   // stn[3].wipBtn[49,6] := 1000;
   // stn[3].wipBtn[49,7] := 1000;
   // stn[4].wipBtn[0,0] := 1000;
   // stn[4].wipBtn[0,1] := 1000;
   // stn[4].wipBtn[0,2] := 1000;
   // stn[4].wipBtn[0,3] := 1000;
   // stn[4].wipBtn[0,4] := 1000;
   // stn[4].wipBtn[0,5] := 1000;
   // stn[4].wipBtn[0,6] := 1000;
   // stn[4].wipBtn[0,7] := 195000;
   // stn[4].wipBtn[1,0] := 1000;
   // stn[4].wipBtn[1,1] := 1000;
   // stn[4].wipBtn[1,2] := 1000;
   // stn[4].wipBtn[1,3] := 1000;
   // stn[4].wipBtn[1,4] := 1000;
   // stn[4].wipBtn[1,5] := 1000;
   // stn[4].wipBtn[1,6] := 1000;
   // stn[4].wipBtn[1,7] := 1000;
   // stn[4].wipBtn[2,0] := 1000;
   // stn[4].wipBtn[2,1] := 1000;
   // stn[4].wipBtn[2,2] := 1000;
   // stn[4].wipBtn[2,3] := 1000;
   // stn[4].wipBtn[2,4] := 1000;
   // stn[4].wipBtn[2,5] := 1000;
   // stn[4].wipBtn[2,6] := 1000;
   // stn[4].wipBtn[2,7] := 1000;
   // stn[4].wipBtn[3,0] := 1000;
   // stn[4].wipBtn[3,1] := 1000;
   // stn[4].wipBtn[3,2] := 1000;
   // stn[4].wipBtn[3,3] := 1000;
   // stn[4].wipBtn[3,4] := 1000;
   // stn[4].wipBtn[3,5] := 1000;
   // stn[4].wipBtn[3,6] := 1000;
   // stn[4].wipBtn[3,7] := 1000;
   // stn[4].wipBtn[4,0] := 1000;
   // stn[4].wipBtn[4,1] := 1000;
   // stn[4].wipBtn[4,2] := 1000;
   // stn[4].wipBtn[4,3] := 1000;
   // stn[4].wipBtn[4,4] := 1000;
   // stn[4].wipBtn[4,5] := 1000;
   // stn[4].wipBtn[4,6] := 1000;
   // stn[4].wipBtn[4,7] := 1000;
   // stn[4].wipBtn[5,0] := 1000;
   // stn[4].wipBtn[5,1] := 1000;
   // stn[4].wipBtn[5,2] := 1000;
   // stn[4].wipBtn[5,3] := 1000;
   // stn[4].wipBtn[5,4] := 1000;
   // stn[4].wipBtn[5,5] := 1000;
   // stn[4].wipBtn[5,6] := 1000;
   // stn[4].wipBtn[5,7] := 1000;
   // stn[4].wipBtn[6,0] := 1000;
   // stn[4].wipBtn[6,1] := 1000;
   // stn[4].wipBtn[6,2] := 1000;
   // stn[4].wipBtn[6,3] := 1000;
   // stn[4].wipBtn[6,4] := 1000;
   // stn[4].wipBtn[6,5] := 1000;
   // stn[4].wipBtn[6,6] := 1000;
   // stn[4].wipBtn[6,7] := 1000;
   // stn[4].wipBtn[7,0] := 1000;
   // stn[4].wipBtn[7,1] := 1000;
   // stn[4].wipBtn[7,2] := 1000;
   // stn[4].wipBtn[7,3] := 1000;
   // stn[4].wipBtn[7,4] := 1000;
   // stn[4].wipBtn[7,5] := 1000;
   // stn[4].wipBtn[7,6] := 1000;
   // stn[4].wipBtn[7,7] := 1000;
   // stn[4].wipBtn[8,0] := 1000;
   // stn[4].wipBtn[8,1] := 1000;
   // stn[4].wipBtn[8,2] := 1000;
   // stn[4].wipBtn[8,3] := 1000;
   // stn[4].wipBtn[8,4] := 1000;
   // stn[4].wipBtn[8,5] := 1000;
   // stn[4].wipBtn[8,6] := 1000;
   // stn[4].wipBtn[8,7] := 1000;
   // stn[4].wipBtn[9,0] := 1000;
   // stn[4].wipBtn[9,1] := 1000;
   // stn[4].wipBtn[9,2] := 1000;
   // stn[4].wipBtn[9,3] := 1000;
   // stn[4].wipBtn[9,4] := 1000;
   // stn[4].wipBtn[9,5] := 1000;
   // stn[4].wipBtn[9,6] := 1000;
   // stn[4].wipBtn[9,7] := 1000;
   // stn[4].wipBtn[10,0] := 1000;
   // stn[4].wipBtn[10,1] := 1000;
   // stn[4].wipBtn[10,2] := 1000;
   // stn[4].wipBtn[10,3] := 1000;
   // stn[4].wipBtn[10,4] := 1000;
   // stn[4].wipBtn[10,5] := 1000;
   // stn[4].wipBtn[10,6] := 1000;
   // stn[4].wipBtn[10,7] := 1000;
   // stn[4].wipBtn[11,0] := 1000;
   // stn[4].wipBtn[11,1] := 1000;
   // stn[4].wipBtn[11,2] := 1000;
   // stn[4].wipBtn[11,3] := 1000;
   // stn[4].wipBtn[11,4] := 1000;
   // stn[4].wipBtn[11,5] := 1000;
   // stn[4].wipBtn[11,6] := 1000;
   // stn[4].wipBtn[11,7] := 1000;
   // stn[4].wipBtn[12,0] := 1000;
   // stn[4].wipBtn[12,1] := 1000;
   // stn[4].wipBtn[12,2] := 1000;
   // stn[4].wipBtn[12,3] := 1000;
   // stn[4].wipBtn[12,4] := 1000;
   // stn[4].wipBtn[12,5] := 1000;
   // stn[4].wipBtn[12,6] := 1000;
   // stn[4].wipBtn[12,7] := 1000;
   // stn[4].wipBtn[13,0] := 1000;
   // stn[4].wipBtn[13,1] := 1000;
   // stn[4].wipBtn[13,2] := 1000;
   // stn[4].wipBtn[13,3] := 1000;
   // stn[4].wipBtn[13,4] := 1000;
   // stn[4].wipBtn[13,5] := 1000;
   // stn[4].wipBtn[13,6] := 1000;
   // stn[4].wipBtn[13,7] := 1000;
   // stn[4].wipBtn[14,0] := 1000;
   // stn[4].wipBtn[14,1] := 1000;
   // stn[4].wipBtn[14,2] := 1000;
   // stn[4].wipBtn[14,3] := 1000;
   // stn[4].wipBtn[14,4] := 1000;
   // stn[4].wipBtn[14,5] := 1000;
   // stn[4].wipBtn[14,6] := 1000;
   // stn[4].wipBtn[14,7] := 1000;
   // stn[4].wipBtn[15,0] := 1000;
   // stn[4].wipBtn[15,1] := 1000;
   // stn[4].wipBtn[15,2] := 1000;
   // stn[4].wipBtn[15,3] := 1000;
   // stn[4].wipBtn[15,4] := 1000;
   // stn[4].wipBtn[15,5] := 1000;
   // stn[4].wipBtn[15,6] := 1000;
   // stn[4].wipBtn[15,7] := 1000;
   // stn[4].wipBtn[16,0] := 1000;
   // stn[4].wipBtn[16,1] := 1000;
   // stn[4].wipBtn[16,2] := 1000;
   // stn[4].wipBtn[16,3] := 1000;
   // stn[4].wipBtn[16,4] := 1000;
   // stn[4].wipBtn[16,5] := 1000;
   // stn[4].wipBtn[16,6] := 1000;
   // stn[4].wipBtn[16,7] := 1000;
   // stn[4].wipBtn[17,0] := 1000;
   // stn[4].wipBtn[17,1] := 1000;
   // stn[4].wipBtn[17,2] := 1000;
   // stn[4].wipBtn[17,3] := 1000;
   // stn[4].wipBtn[17,4] := 1000;
   // stn[4].wipBtn[17,5] := 1000;
   // stn[4].wipBtn[17,6] := 1000;
   // stn[4].wipBtn[17,7] := 1000;
   // stn[4].wipBtn[18,0] := 1000;
   // stn[4].wipBtn[18,1] := 1000;
   // stn[4].wipBtn[18,2] := 1000;
   // stn[4].wipBtn[18,3] := 1000;
   // stn[4].wipBtn[18,4] := 1000;
   // stn[4].wipBtn[18,5] := 1000;
   // stn[4].wipBtn[18,6] := 1000;
   // stn[4].wipBtn[18,7] := 1000;
   // stn[4].wipBtn[19,0] := 1000;
   // stn[4].wipBtn[19,1] := 1000;
   // stn[4].wipBtn[19,2] := 1000;
   // stn[4].wipBtn[19,3] := 1000;
   // stn[4].wipBtn[19,4] := 1000;
   // stn[4].wipBtn[19,5] := 1000;
   // stn[4].wipBtn[19,6] := 1000;
   // stn[4].wipBtn[19,7] := 1000;
   // stn[4].wipBtn[20,0] := 1000;
   // stn[4].wipBtn[20,1] := 1000;
   // stn[4].wipBtn[20,2] := 1000;
   // stn[4].wipBtn[20,3] := 1000;
   // stn[4].wipBtn[20,4] := 1000;
   // stn[4].wipBtn[20,5] := 1000;
   // stn[4].wipBtn[20,6] := 1000;
   // stn[4].wipBtn[20,7] := 1000;
   // stn[4].wipBtn[21,0] := 1000;
   // stn[4].wipBtn[21,1] := 1000;
   // stn[4].wipBtn[21,2] := 1000;
   // stn[4].wipBtn[21,3] := 1000;
   // stn[4].wipBtn[21,4] := 1000;
   // stn[4].wipBtn[21,5] := 1000;
   // stn[4].wipBtn[21,6] := 1000;
   // stn[4].wipBtn[21,7] := 1000;
   // stn[4].wipBtn[22,0] := 1000;
   // stn[4].wipBtn[22,1] := 1000;
   // stn[4].wipBtn[22,2] := 1000;
   // stn[4].wipBtn[22,3] := 1000;
   // stn[4].wipBtn[22,4] := 1000;
   // stn[4].wipBtn[22,5] := 1000;
   // stn[4].wipBtn[22,6] := 1000;
   // stn[4].wipBtn[22,7] := 1000;
   // stn[4].wipBtn[23,0] := 1000;
   // stn[4].wipBtn[23,1] := 1000;
   // stn[4].wipBtn[23,2] := 1000;
   // stn[4].wipBtn[23,3] := 1000;
   // stn[4].wipBtn[23,4] := 1000;
   // stn[4].wipBtn[23,5] := 1000;
   // stn[4].wipBtn[23,6] := 1000;
   // stn[4].wipBtn[23,7] := 1000;
   // stn[4].wipBtn[24,0] := 1000;
   // stn[4].wipBtn[24,1] := 1000;
   // stn[4].wipBtn[24,2] := 1000;
   // stn[4].wipBtn[24,3] := 1000;
   // stn[4].wipBtn[24,4] := 1000;
   // stn[4].wipBtn[24,5] := 1000;
   // stn[4].wipBtn[24,6] := 1000;
   // stn[4].wipBtn[24,7] := 1000;
   // stn[4].wipBtn[25,0] := 1000;
   // stn[4].wipBtn[25,1] := 1000;
   // stn[4].wipBtn[25,2] := 1000;
   // stn[4].wipBtn[25,3] := 1000;
   // stn[4].wipBtn[25,4] := 1000;
   // stn[4].wipBtn[25,5] := 1000;
   // stn[4].wipBtn[25,6] := 1000;
   // stn[4].wipBtn[25,7] := 1000;
   // stn[4].wipBtn[26,0] := 1000;
   // stn[4].wipBtn[26,1] := 1000;
   // stn[4].wipBtn[26,2] := 1000;
   // stn[4].wipBtn[26,3] := 1000;
   // stn[4].wipBtn[26,4] := 1000;
   // stn[4].wipBtn[26,5] := 1000;
   // stn[4].wipBtn[26,6] := 1000;
   // stn[4].wipBtn[26,7] := 1000;
   // stn[4].wipBtn[27,0] := 1000;
   // stn[4].wipBtn[27,1] := 1000;
   // stn[4].wipBtn[27,2] := 1000;
   // stn[4].wipBtn[27,3] := 1000;
   // stn[4].wipBtn[27,4] := 1000;
   // stn[4].wipBtn[27,5] := 1000;
   // stn[4].wipBtn[27,6] := 1000;
   // stn[4].wipBtn[27,7] := 1000;
   // stn[4].wipBtn[28,0] := 1000;
   // stn[4].wipBtn[28,1] := 1000;
   // stn[4].wipBtn[28,2] := 1000;
   // stn[4].wipBtn[28,3] := 1000;
   // stn[4].wipBtn[28,4] := 1000;
   // stn[4].wipBtn[28,5] := 1000;
   // stn[4].wipBtn[28,6] := 1000;
   // stn[4].wipBtn[28,7] := 1000;
   // stn[4].wipBtn[29,0] := 1000;
   // stn[4].wipBtn[29,1] := 1000;
   // stn[4].wipBtn[29,2] := 1000;
   // stn[4].wipBtn[29,3] := 1000;
   // stn[4].wipBtn[29,4] := 1000;
   // stn[4].wipBtn[29,5] := 1000;
   // stn[4].wipBtn[29,6] := 1000;
   // stn[4].wipBtn[29,7] := 1000;
   // stn[4].wipBtn[30,0] := 1000;
   // stn[4].wipBtn[30,1] := 1000;
   // stn[4].wipBtn[30,2] := 1000;
   // stn[4].wipBtn[30,3] := 1000;
   // stn[4].wipBtn[30,4] := 1000;
   // stn[4].wipBtn[30,5] := 1000;
   // stn[4].wipBtn[30,6] := 1000;
   // stn[4].wipBtn[30,7] := 1000;
   // stn[4].wipBtn[31,0] := 1000;
   // stn[4].wipBtn[31,1] := 1000;
   // stn[4].wipBtn[31,2] := 1000;
   // stn[4].wipBtn[31,3] := 1000;
   // stn[4].wipBtn[31,4] := 1000;
   // stn[4].wipBtn[31,5] := 1000;
   // stn[4].wipBtn[31,6] := 1000;
   // stn[4].wipBtn[31,7] := 1000;
   // stn[4].wipBtn[32,0] := 1000;
   // stn[4].wipBtn[32,1] := 1000;
   // stn[4].wipBtn[32,2] := 1000;
   // stn[4].wipBtn[32,3] := 1000;
   // stn[4].wipBtn[32,4] := 1000;
   // stn[4].wipBtn[32,5] := 1000;
   // stn[4].wipBtn[32,6] := 1000;
   // stn[4].wipBtn[32,7] := 1000;
   // stn[4].wipBtn[33,0] := 1000;
   // stn[4].wipBtn[33,1] := 1000;
   // stn[4].wipBtn[33,2] := 1000;
   // stn[4].wipBtn[33,3] := 1000;
   // stn[4].wipBtn[33,4] := 1000;
   // stn[4].wipBtn[33,5] := 1000;
   // stn[4].wipBtn[33,6] := 1000;
   // stn[4].wipBtn[33,7] := 1000;
   // stn[4].wipBtn[34,0] := 1000;
   // stn[4].wipBtn[34,1] := 1000;
   // stn[4].wipBtn[34,2] := 1000;
   // stn[4].wipBtn[34,3] := 1000;
   // stn[4].wipBtn[34,4] := 1000;
   // stn[4].wipBtn[34,5] := 1000;
   // stn[4].wipBtn[34,6] := 1000;
   // stn[4].wipBtn[34,7] := 1000;
   // stn[4].wipBtn[35,0] := 1000;
   // stn[4].wipBtn[35,1] := 1000;
   // stn[4].wipBtn[35,2] := 1000;
   // stn[4].wipBtn[35,3] := 1000;
   // stn[4].wipBtn[35,4] := 1000;
   // stn[4].wipBtn[35,5] := 1000;
   // stn[4].wipBtn[35,6] := 1000;
   // stn[4].wipBtn[35,7] := 1000;
   // stn[4].wipBtn[36,0] := 1000;
   // stn[4].wipBtn[36,1] := 1000;
   // stn[4].wipBtn[36,2] := 1000;
   // stn[4].wipBtn[36,3] := 1000;
   // stn[4].wipBtn[36,4] := 1000;
   // stn[4].wipBtn[36,5] := 1000;
   // stn[4].wipBtn[36,6] := 1000;
   // stn[4].wipBtn[36,7] := 1000;
   // stn[4].wipBtn[37,0] := 1000;
   // stn[4].wipBtn[37,1] := 1000;
   // stn[4].wipBtn[37,2] := 1000;
   // stn[4].wipBtn[37,3] := 1000;
   // stn[4].wipBtn[37,4] := 1000;
   // stn[4].wipBtn[37,5] := 1000;
   // stn[4].wipBtn[37,6] := 1000;
   // stn[4].wipBtn[37,7] := 1000;
   // stn[4].wipBtn[38,0] := 1000;
   // stn[4].wipBtn[38,1] := 1000;
   // stn[4].wipBtn[38,2] := 1000;
   // stn[4].wipBtn[38,3] := 1000;
   // stn[4].wipBtn[38,4] := 1000;
   // stn[4].wipBtn[38,5] := 1000;
   // stn[4].wipBtn[38,6] := 1000;
   // stn[4].wipBtn[38,7] := 1000;
   // stn[4].wipBtn[39,0] := 1000;
   // stn[4].wipBtn[39,1] := 1000;
   // stn[4].wipBtn[39,2] := 1000;
   // stn[4].wipBtn[39,3] := 1000;
   // stn[4].wipBtn[39,4] := 1000;
   // stn[4].wipBtn[39,5] := 1000;
   // stn[4].wipBtn[39,6] := 1000;
   // stn[4].wipBtn[39,7] := 1000;
   // stn[4].wipBtn[40,0] := 1000;
   // stn[4].wipBtn[40,1] := 1000;
   // stn[4].wipBtn[40,2] := 1000;
   // stn[4].wipBtn[40,3] := 1000;
   // stn[4].wipBtn[40,4] := 1000;
   // stn[4].wipBtn[40,5] := 1000;
   // stn[4].wipBtn[40,6] := 1000;
   // stn[4].wipBtn[40,7] := 1000;
   // stn[4].wipBtn[41,0] := 1000;
   // stn[4].wipBtn[41,1] := 1000;
   // stn[4].wipBtn[41,2] := 1000;
   // stn[4].wipBtn[41,3] := 1000;
   // stn[4].wipBtn[41,4] := 1000;
   // stn[4].wipBtn[41,5] := 1000;
   // stn[4].wipBtn[41,6] := 1000;
   // stn[4].wipBtn[41,7] := 1000;
   // stn[4].wipBtn[42,0] := 1000;
   // stn[4].wipBtn[42,1] := 1000;
   // stn[4].wipBtn[42,2] := 1000;
   // stn[4].wipBtn[42,3] := 1000;
   // stn[4].wipBtn[42,4] := 1000;
   // stn[4].wipBtn[42,5] := 1000;
   // stn[4].wipBtn[42,6] := 1000;
   // stn[4].wipBtn[42,7] := 1000;
   // stn[4].wipBtn[43,0] := 1000;
   // stn[4].wipBtn[43,1] := 1000;
   // stn[4].wipBtn[43,2] := 1000;
   // stn[4].wipBtn[43,3] := 1000;
   // stn[4].wipBtn[43,4] := 1000;
   // stn[4].wipBtn[43,5] := 1000;
   // stn[4].wipBtn[43,6] := 1000;
   // stn[4].wipBtn[43,7] := 1000;
   // stn[4].wipBtn[44,0] := 1000;
   // stn[4].wipBtn[44,1] := 1000;
   // stn[4].wipBtn[44,2] := 1000;
   // stn[4].wipBtn[44,3] := 1000;
   // stn[4].wipBtn[44,4] := 1000;
   // stn[4].wipBtn[44,5] := 1000;
   // stn[4].wipBtn[44,6] := 1000;
   // stn[4].wipBtn[44,7] := 1000;
   // stn[4].wipBtn[45,0] := 1000;
   // stn[4].wipBtn[45,1] := 1000;
   // stn[4].wipBtn[45,2] := 1000;
   // stn[4].wipBtn[45,3] := 1000;
   // stn[4].wipBtn[45,4] := 1000;
   // stn[4].wipBtn[45,5] := 1000;
   // stn[4].wipBtn[45,6] := 1000;
   // stn[4].wipBtn[45,7] := 1000;
   // stn[4].wipBtn[46,0] := 1000;
   // stn[4].wipBtn[46,1] := 1000;
   // stn[4].wipBtn[46,2] := 1000;
   // stn[4].wipBtn[46,3] := 1000;
   // stn[4].wipBtn[46,4] := 1000;
   // stn[4].wipBtn[46,5] := 1000;
   // stn[4].wipBtn[46,6] := 1000;
   // stn[4].wipBtn[46,7] := 1000;
   // stn[4].wipBtn[47,0] := 1000;
   // stn[4].wipBtn[47,1] := 1000;
   // stn[4].wipBtn[47,2] := 1000;
   // stn[4].wipBtn[47,3] := 1000;
   // stn[4].wipBtn[47,4] := 1000;
   // stn[4].wipBtn[47,5] := 1000;
   // stn[4].wipBtn[47,6] := 1000;
   // stn[4].wipBtn[47,7] := 1000;
   // stn[4].wipBtn[48,0] := 1000;
   // stn[4].wipBtn[48,1] := 1000;
   // stn[4].wipBtn[48,2] := 1000;
   // stn[4].wipBtn[48,3] := 1000;
   // stn[4].wipBtn[48,4] := 1000;
   // stn[4].wipBtn[48,5] := 1000;
   // stn[4].wipBtn[48,6] := 1000;
   // stn[4].wipBtn[48,7] := 1000;
   // stn[4].wipBtn[49,0] := 1000;
   // stn[4].wipBtn[49,1] := 1000;
   // stn[4].wipBtn[49,2] := 1000;
   // stn[4].wipBtn[49,3] := 1000;
   // stn[4].wipBtn[49,4] := 1000;
   // stn[4].wipBtn[49,5] := 1000;
   // stn[4].wipBtn[49,6] := 1000;
   // stn[4].wipBtn[49,7] := 1000;
   // stn[5].wipBtn[0,0] := 1000;
   // stn[5].wipBtn[0,1] := 194000;
   // stn[5].wipBtn[0,2] := 196000;
   // stn[5].wipBtn[0,3] := 177000;
   // stn[5].wipBtn[0,4] := 1000;
   // stn[5].wipBtn[0,5] := 197000;
   // stn[5].wipBtn[0,6] := 178000;
   // stn[5].wipBtn[0,7] := 176000;
   // stn[5].wipBtn[1,0] := 1000;
   // stn[5].wipBtn[1,1] := 1000;
   // stn[5].wipBtn[1,2] := 1000;
   // stn[5].wipBtn[1,3] := 1000;
   // stn[5].wipBtn[1,4] := 1000;
   // stn[5].wipBtn[1,5] := 1000;
   // stn[5].wipBtn[1,6] := 1000;
   // stn[5].wipBtn[1,7] := 1000;
   // stn[5].wipBtn[2,0] := 1000;
   // stn[5].wipBtn[2,1] := 1000;
   // stn[5].wipBtn[2,2] := 1000;
   // stn[5].wipBtn[2,3] := 1000;
   // stn[5].wipBtn[2,4] := 1000;
   // stn[5].wipBtn[2,5] := 1000;
   // stn[5].wipBtn[2,6] := 1000;
   // stn[5].wipBtn[2,7] := 1000;
   // stn[5].wipBtn[3,0] := 1000;
   // stn[5].wipBtn[3,1] := 1000;
   // stn[5].wipBtn[3,2] := 1000;
   // stn[5].wipBtn[3,3] := 1000;
   // stn[5].wipBtn[3,4] := 1000;
   // stn[5].wipBtn[3,5] := 1000;
   // stn[5].wipBtn[3,6] := 1000;
   // stn[5].wipBtn[3,7] := 1000;
   // stn[5].wipBtn[4,0] := 1000;
   // stn[5].wipBtn[4,1] := 1000;
   // stn[5].wipBtn[4,2] := 1000;
   // stn[5].wipBtn[4,3] := 1000;
   // stn[5].wipBtn[4,4] := 1000;
   // stn[5].wipBtn[4,5] := 1000;
   // stn[5].wipBtn[4,6] := 1000;
   // stn[5].wipBtn[4,7] := 1000;
   // stn[5].wipBtn[5,0] := 1000;
   // stn[5].wipBtn[5,1] := 1000;
   // stn[5].wipBtn[5,2] := 1000;
   // stn[5].wipBtn[5,3] := 1000;
   // stn[5].wipBtn[5,4] := 1000;
   // stn[5].wipBtn[5,5] := 1000;
   // stn[5].wipBtn[5,6] := 1000;
   // stn[5].wipBtn[5,7] := 1000;
   // stn[5].wipBtn[6,0] := 1000;
   // stn[5].wipBtn[6,1] := 1000;
   // stn[5].wipBtn[6,2] := 1000;
   // stn[5].wipBtn[6,3] := 1000;
   // stn[5].wipBtn[6,4] := 1000;
   // stn[5].wipBtn[6,5] := 1000;
   // stn[5].wipBtn[6,6] := 1000;
   // stn[5].wipBtn[6,7] := 1000;
   // stn[5].wipBtn[7,0] := 1000;
   // stn[5].wipBtn[7,1] := 1000;
   // stn[5].wipBtn[7,2] := 1000;
   // stn[5].wipBtn[7,3] := 1000;
   // stn[5].wipBtn[7,4] := 1000;
   // stn[5].wipBtn[7,5] := 1000;
   // stn[5].wipBtn[7,6] := 1000;
   // stn[5].wipBtn[7,7] := 1000;
   // stn[5].wipBtn[8,0] := 1000;
   // stn[5].wipBtn[8,1] := 1000;
   // stn[5].wipBtn[8,2] := 1000;
   // stn[5].wipBtn[8,3] := 1000;
   // stn[5].wipBtn[8,4] := 1000;
   // stn[5].wipBtn[8,5] := 1000;
   // stn[5].wipBtn[8,6] := 1000;
   // stn[5].wipBtn[8,7] := 1000;
   // stn[5].wipBtn[9,0] := 1000;
   // stn[5].wipBtn[9,1] := 1000;
   // stn[5].wipBtn[9,2] := 1000;
   // stn[5].wipBtn[9,3] := 1000;
   // stn[5].wipBtn[9,4] := 1000;
   // stn[5].wipBtn[9,5] := 1000;
   // stn[5].wipBtn[9,6] := 1000;
   // stn[5].wipBtn[9,7] := 1000;
   // stn[5].wipBtn[10,0] := 1000;
   // stn[5].wipBtn[10,1] := 1000;
   // stn[5].wipBtn[10,2] := 1000;
   // stn[5].wipBtn[10,3] := 1000;
   // stn[5].wipBtn[10,4] := 1000;
   // stn[5].wipBtn[10,5] := 1000;
   // stn[5].wipBtn[10,6] := 1000;
   // stn[5].wipBtn[10,7] := 1000;
   // stn[5].wipBtn[11,0] := 1000;
   // stn[5].wipBtn[11,1] := 1000;
   // stn[5].wipBtn[11,2] := 1000;
   // stn[5].wipBtn[11,3] := 1000;
   // stn[5].wipBtn[11,4] := 1000;
   // stn[5].wipBtn[11,5] := 1000;
   // stn[5].wipBtn[11,6] := 1000;
   // stn[5].wipBtn[11,7] := 1000;
   // stn[5].wipBtn[12,0] := 1000;
   // stn[5].wipBtn[12,1] := 1000;
   // stn[5].wipBtn[12,2] := 1000;
   // stn[5].wipBtn[12,3] := 1000;
   // stn[5].wipBtn[12,4] := 1000;
   // stn[5].wipBtn[12,5] := 1000;
   // stn[5].wipBtn[12,6] := 1000;
   // stn[5].wipBtn[12,7] := 1000;
   // stn[5].wipBtn[13,0] := 1000;
   // stn[5].wipBtn[13,1] := 1000;
   // stn[5].wipBtn[13,2] := 1000;
   // stn[5].wipBtn[13,3] := 1000;
   // stn[5].wipBtn[13,4] := 1000;
   // stn[5].wipBtn[13,5] := 1000;
   // stn[5].wipBtn[13,6] := 1000;
   // stn[5].wipBtn[13,7] := 1000;
   // stn[5].wipBtn[14,0] := 1000;
   // stn[5].wipBtn[14,1] := 1000;
   // stn[5].wipBtn[14,2] := 1000;
   // stn[5].wipBtn[14,3] := 1000;
   // stn[5].wipBtn[14,4] := 1000;
   // stn[5].wipBtn[14,5] := 1000;
   // stn[5].wipBtn[14,6] := 1000;
   // stn[5].wipBtn[14,7] := 1000;
   // stn[5].wipBtn[15,0] := 1000;
   // stn[5].wipBtn[15,1] := 1000;
   // stn[5].wipBtn[15,2] := 1000;
   // stn[5].wipBtn[15,3] := 1000;
   // stn[5].wipBtn[15,4] := 1000;
   // stn[5].wipBtn[15,5] := 1000;
   // stn[5].wipBtn[15,6] := 1000;
   // stn[5].wipBtn[15,7] := 1000;
   // stn[5].wipBtn[16,0] := 1000;
   // stn[5].wipBtn[16,1] := 1000;
   // stn[5].wipBtn[16,2] := 1000;
   // stn[5].wipBtn[16,3] := 1000;
   // stn[5].wipBtn[16,4] := 1000;
   // stn[5].wipBtn[16,5] := 1000;
   // stn[5].wipBtn[16,6] := 1000;
   // stn[5].wipBtn[16,7] := 1000;
   // stn[5].wipBtn[17,0] := 1000;
   // stn[5].wipBtn[17,1] := 1000;
   // stn[5].wipBtn[17,2] := 1000;
   // stn[5].wipBtn[17,3] := 1000;
   // stn[5].wipBtn[17,4] := 1000;
   // stn[5].wipBtn[17,5] := 1000;
   // stn[5].wipBtn[17,6] := 1000;
   // stn[5].wipBtn[17,7] := 1000;
   // stn[5].wipBtn[18,0] := 1000;
   // stn[5].wipBtn[18,1] := 1000;
   // stn[5].wipBtn[18,2] := 1000;
   // stn[5].wipBtn[18,3] := 1000;
   // stn[5].wipBtn[18,4] := 1000;
   // stn[5].wipBtn[18,5] := 1000;
   // stn[5].wipBtn[18,6] := 1000;
   // stn[5].wipBtn[18,7] := 1000;
   // stn[5].wipBtn[19,0] := 1000;
   // stn[5].wipBtn[19,1] := 1000;
   // stn[5].wipBtn[19,2] := 1000;
   // stn[5].wipBtn[19,3] := 1000;
   // stn[5].wipBtn[19,4] := 1000;
   // stn[5].wipBtn[19,5] := 1000;
   // stn[5].wipBtn[19,6] := 1000;
   // stn[5].wipBtn[19,7] := 1000;
   // stn[5].wipBtn[20,0] := 1000;
   // stn[5].wipBtn[20,1] := 1000;
   // stn[5].wipBtn[20,2] := 1000;
   // stn[5].wipBtn[20,3] := 1000;
   // stn[5].wipBtn[20,4] := 1000;
   // stn[5].wipBtn[20,5] := 1000;
   // stn[5].wipBtn[20,6] := 1000;
   // stn[5].wipBtn[20,7] := 1000;
   // stn[5].wipBtn[21,0] := 1000;
   // stn[5].wipBtn[21,1] := 1000;
   // stn[5].wipBtn[21,2] := 1000;
   // stn[5].wipBtn[21,3] := 1000;
   // stn[5].wipBtn[21,4] := 1000;
   // stn[5].wipBtn[21,5] := 1000;
   // stn[5].wipBtn[21,6] := 1000;
   // stn[5].wipBtn[21,7] := 1000;
   // stn[5].wipBtn[22,0] := 1000;
   // stn[5].wipBtn[22,1] := 1000;
   // stn[5].wipBtn[22,2] := 1000;
   // stn[5].wipBtn[22,3] := 1000;
   // stn[5].wipBtn[22,4] := 1000;
   // stn[5].wipBtn[22,5] := 1000;
   // stn[5].wipBtn[22,6] := 1000;
   // stn[5].wipBtn[22,7] := 1000;
   // stn[5].wipBtn[23,0] := 1000;
   // stn[5].wipBtn[23,1] := 1000;
   // stn[5].wipBtn[23,2] := 1000;
   // stn[5].wipBtn[23,3] := 1000;
   // stn[5].wipBtn[23,4] := 1000;
   // stn[5].wipBtn[23,5] := 1000;
   // stn[5].wipBtn[23,6] := 1000;
   // stn[5].wipBtn[23,7] := 1000;
   // stn[5].wipBtn[24,0] := 1000;
   // stn[5].wipBtn[24,1] := 1000;
   // stn[5].wipBtn[24,2] := 1000;
   // stn[5].wipBtn[24,3] := 1000;
   // stn[5].wipBtn[24,4] := 1000;
   // stn[5].wipBtn[24,5] := 1000;
   // stn[5].wipBtn[24,6] := 1000;
   // stn[5].wipBtn[24,7] := 1000;
   // stn[5].wipBtn[25,0] := 1000;
   // stn[5].wipBtn[25,1] := 1000;
   // stn[5].wipBtn[25,2] := 1000;
   // stn[5].wipBtn[25,3] := 1000;
   // stn[5].wipBtn[25,4] := 1000;
   // stn[5].wipBtn[25,5] := 1000;
   // stn[5].wipBtn[25,6] := 1000;
   // stn[5].wipBtn[25,7] := 1000;
   // stn[5].wipBtn[26,0] := 1000;
   // stn[5].wipBtn[26,1] := 1000;
   // stn[5].wipBtn[26,2] := 1000;
   // stn[5].wipBtn[26,3] := 1000;
   // stn[5].wipBtn[26,4] := 1000;
   // stn[5].wipBtn[26,5] := 1000;
   // stn[5].wipBtn[26,6] := 1000;
   // stn[5].wipBtn[26,7] := 1000;
   // stn[5].wipBtn[27,0] := 1000;
   // stn[5].wipBtn[27,1] := 1000;
   // stn[5].wipBtn[27,2] := 1000;
   // stn[5].wipBtn[27,3] := 1000;
   // stn[5].wipBtn[27,4] := 1000;
   // stn[5].wipBtn[27,5] := 1000;
   // stn[5].wipBtn[27,6] := 1000;
   // stn[5].wipBtn[27,7] := 1000;
   // stn[5].wipBtn[28,0] := 1000;
   // stn[5].wipBtn[28,1] := 1000;
   // stn[5].wipBtn[28,2] := 1000;
   // stn[5].wipBtn[28,3] := 1000;
   // stn[5].wipBtn[28,4] := 1000;
   // stn[5].wipBtn[28,5] := 1000;
   // stn[5].wipBtn[28,6] := 1000;
   // stn[5].wipBtn[28,7] := 1000;
   // stn[5].wipBtn[29,0] := 1000;
   // stn[5].wipBtn[29,1] := 1000;
   // stn[5].wipBtn[29,2] := 1000;
   // stn[5].wipBtn[29,3] := 1000;
   // stn[5].wipBtn[29,4] := 1000;
   // stn[5].wipBtn[29,5] := 1000;
   // stn[5].wipBtn[29,6] := 1000;
   // stn[5].wipBtn[29,7] := 1000;
   // stn[5].wipBtn[30,0] := 1000;
   // stn[5].wipBtn[30,1] := 1000;
   // stn[5].wipBtn[30,2] := 1000;
   // stn[5].wipBtn[30,3] := 1000;
   // stn[5].wipBtn[30,4] := 1000;
   // stn[5].wipBtn[30,5] := 1000;
   // stn[5].wipBtn[30,6] := 1000;
   // stn[5].wipBtn[30,7] := 1000;
   // stn[5].wipBtn[31,0] := 1000;
   // stn[5].wipBtn[31,1] := 1000;
   // stn[5].wipBtn[31,2] := 1000;
   // stn[5].wipBtn[31,3] := 1000;
   // stn[5].wipBtn[31,4] := 1000;
   // stn[5].wipBtn[31,5] := 1000;
   // stn[5].wipBtn[31,6] := 1000;
   // stn[5].wipBtn[31,7] := 1000;
   // stn[5].wipBtn[32,0] := 1000;
   // stn[5].wipBtn[32,1] := 1000;
   // stn[5].wipBtn[32,2] := 1000;
   // stn[5].wipBtn[32,3] := 1000;
   // stn[5].wipBtn[32,4] := 1000;
   // stn[5].wipBtn[32,5] := 1000;
   // stn[5].wipBtn[32,6] := 1000;
   // stn[5].wipBtn[32,7] := 1000;
   // stn[5].wipBtn[33,0] := 1000;
   // stn[5].wipBtn[33,1] := 1000;
   // stn[5].wipBtn[33,2] := 1000;
   // stn[5].wipBtn[33,3] := 1000;
   // stn[5].wipBtn[33,4] := 1000;
   // stn[5].wipBtn[33,5] := 1000;
   // stn[5].wipBtn[33,6] := 1000;
   // stn[5].wipBtn[33,7] := 1000;
   // stn[5].wipBtn[34,0] := 1000;
   // stn[5].wipBtn[34,1] := 1000;
   // stn[5].wipBtn[34,2] := 1000;
   // stn[5].wipBtn[34,3] := 1000;
   // stn[5].wipBtn[34,4] := 1000;
   // stn[5].wipBtn[34,5] := 1000;
   // stn[5].wipBtn[34,6] := 1000;
   // stn[5].wipBtn[34,7] := 1000;
   // stn[5].wipBtn[35,0] := 1000;
   // stn[5].wipBtn[35,1] := 1000;
   // stn[5].wipBtn[35,2] := 1000;
   // stn[5].wipBtn[35,3] := 1000;
   // stn[5].wipBtn[35,4] := 1000;
   // stn[5].wipBtn[35,5] := 1000;
   // stn[5].wipBtn[35,6] := 1000;
   // stn[5].wipBtn[35,7] := 1000;
   // stn[5].wipBtn[36,0] := 1000;
   // stn[5].wipBtn[36,1] := 1000;
   // stn[5].wipBtn[36,2] := 1000;
   // stn[5].wipBtn[36,3] := 1000;
   // stn[5].wipBtn[36,4] := 1000;
   // stn[5].wipBtn[36,5] := 1000;
   // stn[5].wipBtn[36,6] := 1000;
   // stn[5].wipBtn[36,7] := 1000;
   // stn[5].wipBtn[37,0] := 1000;
   // stn[5].wipBtn[37,1] := 1000;
   // stn[5].wipBtn[37,2] := 1000;
   // stn[5].wipBtn[37,3] := 1000;
   // stn[5].wipBtn[37,4] := 1000;
   // stn[5].wipBtn[37,5] := 1000;
   // stn[5].wipBtn[37,6] := 1000;
   // stn[5].wipBtn[37,7] := 1000;
   // stn[5].wipBtn[38,0] := 1000;
   // stn[5].wipBtn[38,1] := 1000;
   // stn[5].wipBtn[38,2] := 1000;
   // stn[5].wipBtn[38,3] := 1000;
   // stn[5].wipBtn[38,4] := 1000;
   // stn[5].wipBtn[38,5] := 1000;
   // stn[5].wipBtn[38,6] := 1000;
   // stn[5].wipBtn[38,7] := 1000;
   // stn[5].wipBtn[39,0] := 1000;
   // stn[5].wipBtn[39,1] := 1000;
   // stn[5].wipBtn[39,2] := 1000;
   // stn[5].wipBtn[39,3] := 1000;
   // stn[5].wipBtn[39,4] := 1000;
   // stn[5].wipBtn[39,5] := 1000;
   // stn[5].wipBtn[39,6] := 1000;
   // stn[5].wipBtn[39,7] := 1000;
   // stn[5].wipBtn[40,0] := 1000;
   // stn[5].wipBtn[40,1] := 1000;
   // stn[5].wipBtn[40,2] := 1000;
   // stn[5].wipBtn[40,3] := 1000;
   // stn[5].wipBtn[40,4] := 1000;
   // stn[5].wipBtn[40,5] := 1000;
   // stn[5].wipBtn[40,6] := 1000;
   // stn[5].wipBtn[40,7] := 1000;
   // stn[5].wipBtn[41,0] := 1000;
   // stn[5].wipBtn[41,1] := 1000;
   // stn[5].wipBtn[41,2] := 1000;
   // stn[5].wipBtn[41,3] := 1000;
   // stn[5].wipBtn[41,4] := 1000;
   // stn[5].wipBtn[41,5] := 1000;
   // stn[5].wipBtn[41,6] := 1000;
   // stn[5].wipBtn[41,7] := 1000;
   // stn[5].wipBtn[42,0] := 1000;
   // stn[5].wipBtn[42,1] := 1000;
   // stn[5].wipBtn[42,2] := 1000;
   // stn[5].wipBtn[42,3] := 1000;
   // stn[5].wipBtn[42,4] := 1000;
   // stn[5].wipBtn[42,5] := 1000;
   // stn[5].wipBtn[42,6] := 1000;
   // stn[5].wipBtn[42,7] := 1000;
   // stn[5].wipBtn[43,0] := 1000;
   // stn[5].wipBtn[43,1] := 1000;
   // stn[5].wipBtn[43,2] := 1000;
   // stn[5].wipBtn[43,3] := 1000;
   // stn[5].wipBtn[43,4] := 1000;
   // stn[5].wipBtn[43,5] := 1000;
   // stn[5].wipBtn[43,6] := 1000;
   // stn[5].wipBtn[43,7] := 1000;
   // stn[5].wipBtn[44,0] := 1000;
   // stn[5].wipBtn[44,1] := 1000;
   // stn[5].wipBtn[44,2] := 1000;
   // stn[5].wipBtn[44,3] := 1000;
   // stn[5].wipBtn[44,4] := 1000;
   // stn[5].wipBtn[44,5] := 1000;
   // stn[5].wipBtn[44,6] := 1000;
   // stn[5].wipBtn[44,7] := 1000;
   // stn[5].wipBtn[45,0] := 1000;
   // stn[5].wipBtn[45,1] := 1000;
   // stn[5].wipBtn[45,2] := 1000;
   // stn[5].wipBtn[45,3] := 1000;
   // stn[5].wipBtn[45,4] := 1000;
   // stn[5].wipBtn[45,5] := 1000;
   // stn[5].wipBtn[45,6] := 1000;
   // stn[5].wipBtn[45,7] := 1000;
   // stn[5].wipBtn[46,0] := 1000;
   // stn[5].wipBtn[46,1] := 1000;
   // stn[5].wipBtn[46,2] := 1000;
   // stn[5].wipBtn[46,3] := 1000;
   // stn[5].wipBtn[46,4] := 1000;
   // stn[5].wipBtn[46,5] := 1000;
   // stn[5].wipBtn[46,6] := 1000;
   // stn[5].wipBtn[46,7] := 1000;
   // stn[5].wipBtn[47,0] := 1000;
   // stn[5].wipBtn[47,1] := 1000;
   // stn[5].wipBtn[47,2] := 1000;
   // stn[5].wipBtn[47,3] := 1000;
   // stn[5].wipBtn[47,4] := 1000;
   // stn[5].wipBtn[47,5] := 1000;
   // stn[5].wipBtn[47,6] := 1000;
   // stn[5].wipBtn[47,7] := 1000;
   // stn[5].wipBtn[48,0] := 1000;
   // stn[5].wipBtn[48,1] := 1000;
   // stn[5].wipBtn[48,2] := 1000;
   // stn[5].wipBtn[48,3] := 1000;
   // stn[5].wipBtn[48,4] := 1000;
   // stn[5].wipBtn[48,5] := 1000;
   // stn[5].wipBtn[48,6] := 1000;
   // stn[5].wipBtn[48,7] := 1000;
   // stn[5].wipBtn[49,0] := 1000;
   // stn[5].wipBtn[49,1] := 1000;
   // stn[5].wipBtn[49,2] := 1000;
   // stn[5].wipBtn[49,3] := 1000;
   // stn[5].wipBtn[49,4] := 1000;
   // stn[5].wipBtn[49,5] := 1000;
   // stn[5].wipBtn[49,6] := 1000;
   // stn[5].wipBtn[49,7] := 1000;
   // stn[6].wipBtn[0,0] := 1000;
   // stn[6].wipBtn[0,1] := 209000;
   // stn[6].wipBtn[0,2] := 208000;
   // stn[6].wipBtn[0,3] := 211000;
   // stn[6].wipBtn[0,4] := 1000;
   // stn[6].wipBtn[0,5] := 212000;
   // stn[6].wipBtn[0,6] := 207000;
   // stn[6].wipBtn[0,7] := 206000;
   // stn[6].wipBtn[1,0] := 1000;
   // stn[6].wipBtn[1,1] := 1000;
   // stn[6].wipBtn[1,2] := 1000;
   // stn[6].wipBtn[1,3] := 1000;
   // stn[6].wipBtn[1,4] := 1000;
   // stn[6].wipBtn[1,5] := 1000;
   // stn[6].wipBtn[1,6] := 1000;
   // stn[6].wipBtn[1,7] := 1000;
   // stn[6].wipBtn[2,0] := 1000;
   // stn[6].wipBtn[2,1] := 1000;
   // stn[6].wipBtn[2,2] := 1000;
   // stn[6].wipBtn[2,3] := 1000;
   // stn[6].wipBtn[2,4] := 1000;
   // stn[6].wipBtn[2,5] := 1000;
   // stn[6].wipBtn[2,6] := 1000;
   // stn[6].wipBtn[2,7] := 1000;
   // stn[6].wipBtn[3,0] := 1000;
   // stn[6].wipBtn[3,1] := 1000;
   // stn[6].wipBtn[3,2] := 1000;
   // stn[6].wipBtn[3,3] := 1000;
   // stn[6].wipBtn[3,4] := 1000;
   // stn[6].wipBtn[3,5] := 1000;
   // stn[6].wipBtn[3,6] := 1000;
   // stn[6].wipBtn[3,7] := 1000;
   // stn[6].wipBtn[4,0] := 1000;
   // stn[6].wipBtn[4,1] := 1000;
   // stn[6].wipBtn[4,2] := 1000;
   // stn[6].wipBtn[4,3] := 1000;
   // stn[6].wipBtn[4,4] := 1000;
   // stn[6].wipBtn[4,5] := 1000;
   // stn[6].wipBtn[4,6] := 1000;
   // stn[6].wipBtn[4,7] := 1000;
   // stn[6].wipBtn[5,0] := 1000;
   // stn[6].wipBtn[5,1] := 1000;
   // stn[6].wipBtn[5,2] := 1000;
   // stn[6].wipBtn[5,3] := 1000;
   // stn[6].wipBtn[5,4] := 1000;
   // stn[6].wipBtn[5,5] := 1000;
   // stn[6].wipBtn[5,6] := 1000;
   // stn[6].wipBtn[5,7] := 1000;
   // stn[6].wipBtn[6,0] := 1000;
   // stn[6].wipBtn[6,1] := 1000;
   // stn[6].wipBtn[6,2] := 1000;
   // stn[6].wipBtn[6,3] := 1000;
   // stn[6].wipBtn[6,4] := 1000;
   // stn[6].wipBtn[6,5] := 1000;
   // stn[6].wipBtn[6,6] := 1000;
   // stn[6].wipBtn[6,7] := 1000;
   // stn[6].wipBtn[7,0] := 1000;
   // stn[6].wipBtn[7,1] := 1000;
   // stn[6].wipBtn[7,2] := 1000;
   // stn[6].wipBtn[7,3] := 1000;
   // stn[6].wipBtn[7,4] := 1000;
   // stn[6].wipBtn[7,5] := 1000;
   // stn[6].wipBtn[7,6] := 1000;
   // stn[6].wipBtn[7,7] := 1000;
   // stn[6].wipBtn[8,0] := 1000;
   // stn[6].wipBtn[8,1] := 1000;
   // stn[6].wipBtn[8,2] := 1000;
   // stn[6].wipBtn[8,3] := 1000;
   // stn[6].wipBtn[8,4] := 1000;
   // stn[6].wipBtn[8,5] := 1000;
   // stn[6].wipBtn[8,6] := 1000;
   // stn[6].wipBtn[8,7] := 1000;
   // stn[6].wipBtn[9,0] := 1000;
   // stn[6].wipBtn[9,1] := 1000;
   // stn[6].wipBtn[9,2] := 1000;
   // stn[6].wipBtn[9,3] := 1000;
   // stn[6].wipBtn[9,4] := 1000;
   // stn[6].wipBtn[9,5] := 1000;
   // stn[6].wipBtn[9,6] := 1000;
   // stn[6].wipBtn[9,7] := 1000;
   // stn[6].wipBtn[10,0] := 1000;
   // stn[6].wipBtn[10,1] := 1000;
   // stn[6].wipBtn[10,2] := 1000;
   // stn[6].wipBtn[10,3] := 1000;
   // stn[6].wipBtn[10,4] := 1000;
   // stn[6].wipBtn[10,5] := 1000;
   // stn[6].wipBtn[10,6] := 1000;
   // stn[6].wipBtn[10,7] := 1000;
   // stn[6].wipBtn[11,0] := 1000;
   // stn[6].wipBtn[11,1] := 1000;
   // stn[6].wipBtn[11,2] := 1000;
   // stn[6].wipBtn[11,3] := 1000;
   // stn[6].wipBtn[11,4] := 1000;
   // stn[6].wipBtn[11,5] := 1000;
   // stn[6].wipBtn[11,6] := 1000;
   // stn[6].wipBtn[11,7] := 1000;
   // stn[6].wipBtn[12,0] := 1000;
   // stn[6].wipBtn[12,1] := 1000;
   // stn[6].wipBtn[12,2] := 1000;
   // stn[6].wipBtn[12,3] := 1000;
   // stn[6].wipBtn[12,4] := 1000;
   // stn[6].wipBtn[12,5] := 1000;
   // stn[6].wipBtn[12,6] := 1000;
   // stn[6].wipBtn[12,7] := 1000;
   // stn[6].wipBtn[13,0] := 1000;
   // stn[6].wipBtn[13,1] := 1000;
   // stn[6].wipBtn[13,2] := 1000;
   // stn[6].wipBtn[13,3] := 1000;
   // stn[6].wipBtn[13,4] := 1000;
   // stn[6].wipBtn[13,5] := 1000;
   // stn[6].wipBtn[13,6] := 1000;
   // stn[6].wipBtn[13,7] := 1000;
   // stn[6].wipBtn[14,0] := 1000;
   // stn[6].wipBtn[14,1] := 1000;
   // stn[6].wipBtn[14,2] := 1000;
   // stn[6].wipBtn[14,3] := 1000;
   // stn[6].wipBtn[14,4] := 1000;
   // stn[6].wipBtn[14,5] := 1000;
   // stn[6].wipBtn[14,6] := 1000;
   // stn[6].wipBtn[14,7] := 1000;
   // stn[6].wipBtn[15,0] := 1000;
   // stn[6].wipBtn[15,1] := 1000;
   // stn[6].wipBtn[15,2] := 1000;
   // stn[6].wipBtn[15,3] := 1000;
   // stn[6].wipBtn[15,4] := 1000;
   // stn[6].wipBtn[15,5] := 1000;
   // stn[6].wipBtn[15,6] := 1000;
   // stn[6].wipBtn[15,7] := 1000;
   // stn[6].wipBtn[16,0] := 1000;
   // stn[6].wipBtn[16,1] := 1000;
   // stn[6].wipBtn[16,2] := 1000;
   // stn[6].wipBtn[16,3] := 1000;
   // stn[6].wipBtn[16,4] := 1000;
   // stn[6].wipBtn[16,5] := 1000;
   // stn[6].wipBtn[16,6] := 1000;
   // stn[6].wipBtn[16,7] := 1000;
   // stn[6].wipBtn[17,0] := 1000;
   // stn[6].wipBtn[17,1] := 1000;
   // stn[6].wipBtn[17,2] := 1000;
   // stn[6].wipBtn[17,3] := 1000;
   // stn[6].wipBtn[17,4] := 1000;
   // stn[6].wipBtn[17,5] := 1000;
   // stn[6].wipBtn[17,6] := 1000;
   // stn[6].wipBtn[17,7] := 1000;
   // stn[6].wipBtn[18,0] := 1000;
   // stn[6].wipBtn[18,1] := 1000;
   // stn[6].wipBtn[18,2] := 1000;
   // stn[6].wipBtn[18,3] := 1000;
   // stn[6].wipBtn[18,4] := 1000;
   // stn[6].wipBtn[18,5] := 1000;
   // stn[6].wipBtn[18,6] := 1000;
   // stn[6].wipBtn[18,7] := 1000;
   // stn[6].wipBtn[19,0] := 1000;
   // stn[6].wipBtn[19,1] := 1000;
   // stn[6].wipBtn[19,2] := 1000;
   // stn[6].wipBtn[19,3] := 1000;
   // stn[6].wipBtn[19,4] := 1000;